// TIA Portal project "Øvelser_2_3_4_5_6_8" (V16)

(* hardware
DEVICE "S7-1200 station_1"  S7-1200 Station
   slot 0: "Rack_0"  S7-1200 Rack  Rack  V1.0
   slot 1: "PLC_1"  CPU 1214C DC/DC/DC  6ES7 214-1AG40-0XB0  V4.4
   slot 3: "AQ 1x12BIT_1"  AQ1 signal board  6ES7 232-4HA30-0XB0  V1.0
DEVICE "HMI_1"  KTP700 Basic PN
   slot 0: "HMI_1"  KTP700 Basic PN  6AV2 123-2GB03-0AX0  16.0.0.0
   slot 1: "HMI_RT_1"  KTP700 Basic PN  6AV2 123-2GB03-0AX0  16.0.0.0
   slot 5: "HMI_1.IE_CP_1"  PROFINET Interface  16.0.0.0
      slot 1: "PROFINET Interface_1"  PROFINET Interface
         slot 1: "Port_1"  Port
*)

// ===== PLC "PLC_1"  CPU 1214C DC/DC/DC =====

VAR_GLOBAL   // PLC tag table "Default tag table"
   "AutoHighCommand" AT %M2.0 : Bool;
   "TestStatus" AT %MW4 : Word;
   "HighCommand" AT %M2.1 : Bool;
   "LowCommand" AT %M2.2 : Bool;
   "SensorLow" AT %M2.4 : Bool;
   "IsHigh" AT %M2.5 : Bool;
   "IsLow" AT %M2.6 : Bool;
   "SensorIn" AT %I0.0 : Bool;
   "SensorOut" AT %I0.1 : Bool;
   "GoOut" AT %Q0.0 : Bool;
   "GoIn" AT %Q0.1 : Bool;
   "SensorUp" AT %I0.3 : Bool;
   "SensorDown" AT %I0.5 : Bool;
   "GoUp" AT %Q0.3 : Bool;
   "GoDown" AT %Q0.2 : Bool;
   "GrabCommand" AT %Q0.4 : Bool;
   "TestCommands" AT %MW0 : Word;
   "SensorHigh" AT %M2.3 : Bool;
   "IsIn" AT %M2.7 : Bool;
   "IsOut" AT %M3.0 : Bool;
   "AutoCommandGoOut" AT %M3.1 : Bool;
   "AutoCommandGoDown" AT %M3.2 : Bool;
   "AutoCommandGrab" AT %M3.3 : Bool;
   "IsUp" AT %M3.4 : Bool;
   "IsDown" AT %M3.5 : Bool;
   "HasGrapped" AT %M3.6 : Bool;
   "HasReleased" AT %M3.7 : Bool;
END_VAR

TYPE "TypeHMI_Commands"
   STRUCT
      Spare0 : Bool;   // (Bit 8), byteswap
      Spare1 : Bool;
      Spare2 : Bool;
      Spare3 : Bool;
      Spare4 : Bool;
      Spare5 : Bool;
      Spare6 : Bool;
      Spare7 : Bool;
      Manual : Bool;   // (Bit 0), byteswap
      Auto : Bool;
      ManualHighCommand : Bool;
      ManualLowCommand : Bool;
      SimulateFeddback : Bool;   // toggle simulation of feedback sensors
      Spare8 : Bool;
      Spare9 : Bool;
      Spare10 : Bool;
   END_STRUCT;
END_TYPE

TYPE "TypeHMI_Status"
   STRUCT
      AlarmToHigh : Bool;
      AlarmToLow : Bool;
      Spare2 : Bool;
      Spare3 : Bool;
      Spare4 : Bool;
      Spare5 : Bool;
      Spare6 : Bool;
      Spare7 : Bool;
      IsManual : Bool;
      IsHigh : Bool;
      IsLow : Bool;
      TransitionToHigh : Bool;
      TransitionToLow : Bool;
      FeedbackSensorLow : Bool;   // Satus, sensor
      FeedbackSensorHigh : Bool;   // Status, sensor
      FeedbackIsSimulated : Bool;
   END_STRUCT;
END_TYPE

DATA_BLOCK "Type_ControlModuleActuator_DB"   // DB1
{ S7_Optimized_Access := 'TRUE' }
VERSION : 0.1
// stored: InstanceOfName Type_ControlModuleActuator
"Type_ControlModuleActuator"
BEGIN
END_DATA_BLOCK

DATA_BLOCK "Type_ControlModuleActuator_DB_1"   // DB2
{ S7_Optimized_Access := 'TRUE' }
VERSION : 0.1
// stored: InstanceOfName Type_ControlModuleActuator
"Type_ControlModuleActuator"
BEGIN
END_DATA_BLOCK

DATA_BLOCK "Type_ControlModuleActuator_DB_2"   // DB3
{ S7_Optimized_Access := 'TRUE' }
VERSION : 0.1
// stored: InstanceOfName Type_ControlModuleActuator
"Type_ControlModuleActuator"
BEGIN
END_DATA_BLOCK

DATA_BLOCK "HMI"   // DB4
{ S7_Optimized_Access := 'TRUE' }
VERSION : 0.1
   VAR
      InOut : Struct
         Command : Word;
         Status : Word;
         StatusInt : Int;
      END_STRUCT;
      UpDown : Struct
         Command : Word;
         Status : Word;
         StatusInt : Int;
      END_STRUCT;
      Grab : Struct
         Command : Word;
         Status : Word;
         StatusInt : Int;
      END_STRUCT;
      TankCalculation : Struct
         CurrentLiguidLevel : Real;   // m
         Radius : Real;   // m
         ConeHight : Real;   // m
         Content : Real;   // m^3
      END_STRUCT;
      Sequence : Struct
         CommandAToB : Bool;
         CommandBToA : Bool;
         Status : Int;
      END_STRUCT;
   END_VAR
BEGIN
END_DATA_BLOCK

DATA_BLOCK "UpDown"   // DB5
{ S7_Optimized_Access := 'TRUE' }
VERSION : 0.1
// stored: InstanceOfName Type_ControlModuleActuator
"Type_ControlModuleActuator"
BEGIN
END_DATA_BLOCK

DATA_BLOCK "Grab"   // DB6
{ S7_Optimized_Access := 'TRUE' }
VERSION : 0.1
// stored: InstanceOfName Type_ControlModuleActuator
"Type_ControlModuleActuator"
BEGIN
END_DATA_BLOCK

DATA_BLOCK "HMI_alarms"   // DB9
{ S7_Optimized_Access := 'TRUE' }
VERSION : 0.1
   VAR
      alarm1 : Bool;
      alarm2 : Bool;
      alarm3 : Bool;
      alarm4 : Bool;
      alarm5 : Bool;
      alarm6 : Bool;
   END_VAR
BEGIN
END_DATA_BLOCK

DATA_BLOCK "Sequence_DB"   // DB10
{ S7_Optimized_Access := 'TRUE' }
VERSION : 0.1
// stored: InstanceOfName Sequence
"Sequence"
BEGIN
END_DATA_BLOCK

// folder: System blocks/Program resources

DATA_BLOCK "IEC_Timer_0_DB"   // DB7
{ S7_Optimized_Access := 'TRUE' }
AUTHOR : Simatic
FAMILY : IEC
NAME : IEC_TMR
VERSION : 1.0
// stored: InstanceOfName IEC_TIMER
"IEC_TIMER"
BEGIN
END_DATA_BLOCK

DATA_BLOCK "IEC_Timer_0_DB_1"   // DB8
{ S7_Optimized_Access := 'TRUE' }
AUTHOR : Simatic
FAMILY : IEC
NAME : IEC_TMR
VERSION : 1.0
// stored: InstanceOfName IEC_TIMER
"IEC_TIMER"
BEGIN
END_DATA_BLOCK

// folder: (top level)

FUNCTION_BLOCK "Type_ControlModuleActuator"   // FB1, LAD
{ S7_Optimized_Access := 'TRUE' }
VERSION : 0.1
   VAR_INPUT
      InHMICommands : Word;
      HMI_Commands AT InHMICommands : "TypeHMI_Commands";
      AutoHighCommand : Bool;
      FeedbackSensorHigh : Bool;
      FeedbackSensorLow : Bool;
      FeedbackTime : Time;
   END_VAR
   VAR_OUTPUT
      OutHMIStatus : Word;
      HMI_Status AT OutHMIStatus : "TypeHMI_Status";
      StatusInt : Int;
      HighCommand : Bool;
      LowCommand : Bool;
      IsHigh : Bool;
      IsLow : Bool;
   END_VAR
   VAR
      Manual : Bool;
      StaticHighCommand : Bool;
      StaticIsSimulated : Bool;
      SimulatedHigh : Bool;
      SimulatedLow : Bool;
      HighAlarmTimer : TON_TIME;
      LowAlarmTimer : TON_TIME;
   END_VAR
BEGIN

REGION Network 1: Manual/Auto
   // controlled by HMI
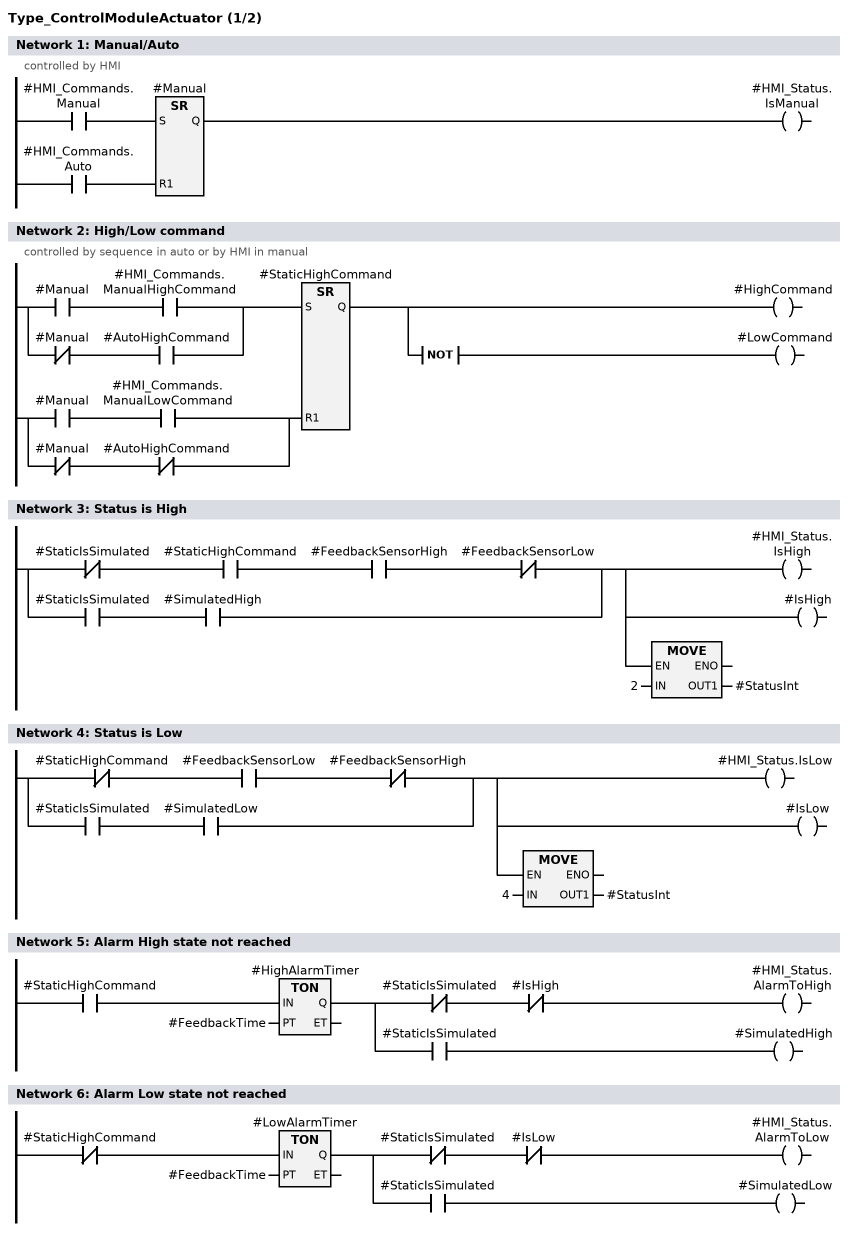
   RUNG wire#powerrail
      Contact( #HMI_Commands.Manual )
      S_SR(operand := #Manual, r1 := wire#w1)
      Coil( #HMI_Status.IsManual )
   END_RUNG
   RUNG wire#powerrail
      Contact( #HMI_Commands.Auto )
   END_RUNG wire#w1
   // the same network as SCL:
   IF #HMI_Commands.Manual THEN
       #Manual := TRUE;   // SR flip-flop
   END_IF;
   IF #HMI_Commands.Auto THEN #Manual := FALSE; END_IF;
   #HMI_Status.IsManual := #Manual;
END_REGION

REGION Network 2: High/Low command
   // controlled by sequence in auto or by HMI in manual
   RUNG wire#powerrail
      Contact( #Manual )
      Contact( #HMI_Commands.ManualHighCommand )
      wire#w1
      S_SR(operand := #StaticHighCommand, r1 := wire#w2)
      wire#w3
      Coil( #HighCommand )
   END_RUNG
   RUNG wire#powerrail
      I_Contact( #Manual )
      Contact( #AutoHighCommand )
   END_RUNG wire#w1
   RUNG wire#powerrail
      Contact( #Manual )
      Contact( #HMI_Commands.ManualLowCommand )
   END_RUNG wire#w2
   RUNG wire#powerrail
      I_Contact( #Manual )
      I_Contact( #AutoHighCommand )
   END_RUNG wire#w2
   RUNG wire#w3
      Not()
      Coil( #LowCommand )
   END_RUNG
   // the same network as SCL:
   IF (#Manual AND #HMI_Commands.ManualHighCommand) OR (NOT #Manual AND #AutoHighCommand) THEN
       #StaticHighCommand := TRUE;   // SR flip-flop
   END_IF;
   IF (#Manual AND #HMI_Commands.ManualLowCommand) OR (NOT #Manual AND NOT #AutoHighCommand) THEN
       #StaticHighCommand := FALSE;
   END_IF;
   #HighCommand := #StaticHighCommand;
   #LowCommand := NOT #StaticHighCommand;
END_REGION

REGION Network 3: Status is High
   RUNG wire#powerrail
      I_Contact( #StaticIsSimulated )
      Contact( #StaticHighCommand )
      Contact( #FeedbackSensorHigh )
      I_Contact( #FeedbackSensorLow )
      wire#w1
      Coil( #HMI_Status.IsHigh )
   END_RUNG
   RUNG wire#powerrail
      Contact( #StaticIsSimulated )
      Contact( #SimulatedHigh )
   END_RUNG wire#w1
   RUNG wire#w1
      Coil( #IsHigh )
   END_RUNG
   RUNG wire#w1
      Move(in := 2, out1 => #StatusInt)
   END_RUNG
   // the same network as SCL:
   #HMI_Status.IsHigh := (NOT #StaticIsSimulated AND #StaticHighCommand AND #FeedbackSensorHigh AND NOT #FeedbackSensorLow) OR (#StaticIsSimulated AND #SimulatedHigh);
   #IsHigh := #HMI_Status.IsHigh;
   IF #HMI_Status.IsHigh THEN #StatusInt := 2; END_IF;
END_REGION

REGION Network 4: Status is Low
   RUNG wire#powerrail
      I_Contact( #StaticHighCommand )
      Contact( #FeedbackSensorLow )
      I_Contact( #FeedbackSensorHigh )
      wire#w1
      Coil( #HMI_Status.IsLow )
   END_RUNG
   RUNG wire#powerrail
      Contact( #StaticIsSimulated )
      Contact( #SimulatedLow )
   END_RUNG wire#w1
   RUNG wire#w1
      Coil( #IsLow )
   END_RUNG
   RUNG wire#w1
      Move(in := 4, out1 => #StatusInt)
   END_RUNG
   // the same network as SCL:
   #HMI_Status.IsLow := (NOT #StaticHighCommand AND #FeedbackSensorLow AND NOT #FeedbackSensorHigh) OR (#StaticIsSimulated AND #SimulatedLow);
   #IsLow := #HMI_Status.IsLow;
   IF #HMI_Status.IsLow THEN #StatusInt := 4; END_IF;
END_REGION

REGION Network 5: Alarm High state not reached
   #HighAlarmTimer(IN := #StaticHighCommand, PT := #FeedbackTime);   // TON
   #HMI_Status.AlarmToHigh := #HighAlarmTimer.Q AND NOT #StaticIsSimulated AND NOT #IsHigh;
   #SimulatedHigh := #HighAlarmTimer.Q AND #StaticIsSimulated;
END_REGION

REGION Network 6: Alarm Low state not reached
   #LowAlarmTimer(IN := NOT #StaticHighCommand, PT := #FeedbackTime);   // TON
   #HMI_Status.AlarmToLow := #LowAlarmTimer.Q AND NOT #StaticIsSimulated AND NOT #IsLow;
   #SimulatedLow := #LowAlarmTimer.Q AND #StaticIsSimulated;
END_REGION

REGION Network 7: Togle simulation
END_REGION

REGION Network 8: Transition to High
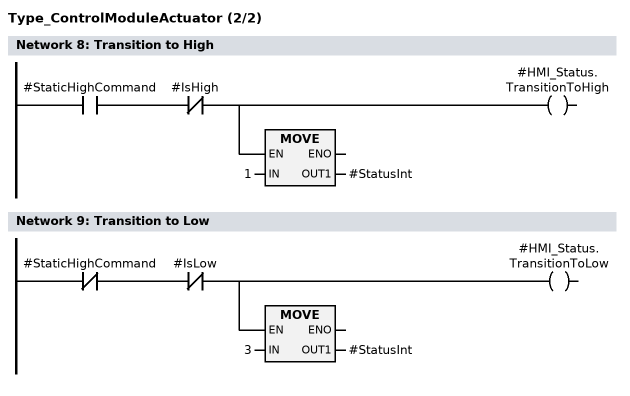
   RUNG wire#powerrail
      Contact( #StaticHighCommand )
      I_Contact( #IsHigh )
      wire#w1
      Coil( #HMI_Status.TransitionToHigh )
   END_RUNG
   RUNG wire#w1
      Move(in := 1, out1 => #StatusInt)
   END_RUNG
   // the same network as SCL:
   #HMI_Status.TransitionToHigh := #StaticHighCommand AND NOT #IsHigh;
   IF #HMI_Status.TransitionToHigh THEN #StatusInt := 1; END_IF;
END_REGION

REGION Network 9: Transition to Low
   RUNG wire#powerrail
      I_Contact( #StaticHighCommand )
      I_Contact( #IsLow )
      wire#w1
      Coil( #HMI_Status.TransitionToLow )
   END_RUNG
   RUNG wire#w1
      Move(in := 3, out1 => #StatusInt)
   END_RUNG
   // the same network as SCL:
   #HMI_Status.TransitionToLow := NOT #StaticHighCommand AND NOT #IsLow;
   IF #HMI_Status.TransitionToLow THEN #StatusInt := 3; END_IF;
END_REGION
END_FUNCTION_BLOCK

FUNCTION_BLOCK "Sequence"   // FB2, LAD
{ S7_Optimized_Access := 'TRUE' }
VERSION : 0.1
   VAR_INPUT
      AToB : Bool;
      BtoA : Bool;
      IsIn : Bool;
      IsOut : Bool;
      IsUp : Bool;
      IsDown : Bool;
      HasGrapped : Bool;
      HasReleased : Bool;
   END_VAR
   VAR_OUTPUT
      AutoCommandGoOut : Bool;
      AutoCommandGoDown : Bool;
      AutoCommandGrab : Bool;
      StatusStepNr : Int;
   END_VAR
   VAR
      StepNr : Int;
   END_VAR
   VAR_TEMP   // added for the SCL form of the ladder/FBD networks
      _w1 : Bool;
   END_VAR
BEGIN

REGION Network 1: Step 0:Idle
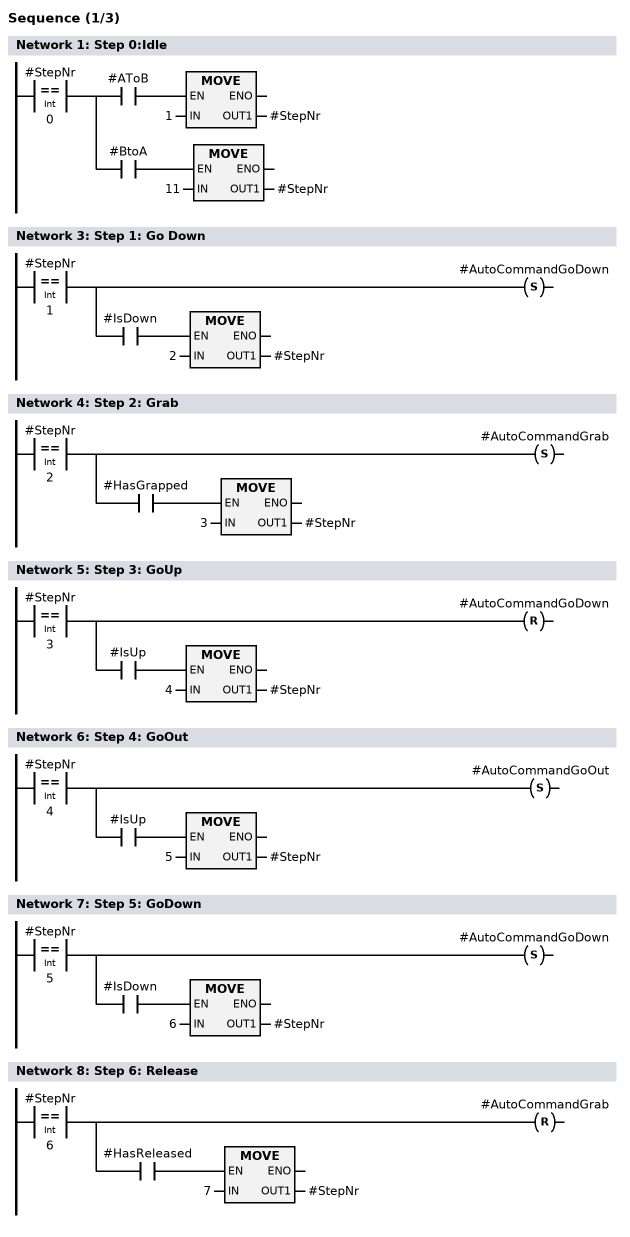
   RUNG wire#powerrail
      { S7_Templates := "SrcType := Int" } EQ_Contact(in1 := #StepNr, in2 := 0)
      wire#w1
      Contact( #AToB )
      Move(in := 1, out1 => #StepNr)
   END_RUNG
   RUNG wire#w1
      Contact( #BtoA )
      Move(in := 11, out1 => #StepNr)
   END_RUNG
   // the same network as SCL:
   #_w1 := #StepNr = 0;
   IF #_w1 AND #AToB THEN #StepNr := 1; END_IF;
   IF #_w1 AND #BtoA THEN #StepNr := 11; END_IF;
END_REGION

REGION Network 2: AToB
END_REGION

REGION Network 3: Step 1: Go Down
   RUNG wire#powerrail
      { S7_Templates := "SrcType := Int" } EQ_Contact(in1 := #StepNr, in2 := 1)
      wire#w1
      S_Coil( #AutoCommandGoDown )
   END_RUNG
   RUNG wire#w1
      Contact( #IsDown )
      Move(in := 2, out1 => #StepNr)
   END_RUNG
   // the same network as SCL:
   #_w1 := #StepNr = 1;
   IF #_w1 THEN #AutoCommandGoDown := TRUE; END_IF;
   IF #_w1 AND #IsDown THEN #StepNr := 2; END_IF;
END_REGION

REGION Network 4: Step 2: Grab
   RUNG wire#powerrail
      { S7_Templates := "SrcType := Int" } EQ_Contact(in1 := #StepNr, in2 := 2)
      wire#w1
      S_Coil( #AutoCommandGrab )
   END_RUNG
   RUNG wire#w1
      Contact( #HasGrapped )
      Move(in := 3, out1 => #StepNr)
   END_RUNG
   // the same network as SCL:
   #_w1 := #StepNr = 2;
   IF #_w1 THEN #AutoCommandGrab := TRUE; END_IF;
   IF #_w1 AND #HasGrapped THEN #StepNr := 3; END_IF;
END_REGION

REGION Network 5: Step 3: GoUp
   RUNG wire#powerrail
      { S7_Templates := "SrcType := Int" } EQ_Contact(in1 := #StepNr, in2 := 3)
      wire#w1
      R_Coil( #AutoCommandGoDown )
   END_RUNG
   RUNG wire#w1
      Contact( #IsUp )
      Move(in := 4, out1 => #StepNr)
   END_RUNG
   // the same network as SCL:
   #_w1 := #StepNr = 3;
   IF #_w1 THEN #AutoCommandGoDown := FALSE; END_IF;
   IF #_w1 AND #IsUp THEN #StepNr := 4; END_IF;
END_REGION

REGION Network 6: Step 4: GoOut
   RUNG wire#powerrail
      { S7_Templates := "SrcType := Int" } EQ_Contact(in1 := #StepNr, in2 := 4)
      wire#w1
      S_Coil( #AutoCommandGoOut )
   END_RUNG
   RUNG wire#w1
      Contact( #IsUp )
      Move(in := 5, out1 => #StepNr)
   END_RUNG
   // the same network as SCL:
   #_w1 := #StepNr = 4;
   IF #_w1 THEN #AutoCommandGoOut := TRUE; END_IF;
   IF #_w1 AND #IsUp THEN #StepNr := 5; END_IF;
END_REGION

REGION Network 7: Step 5: GoDown
   RUNG wire#powerrail
      { S7_Templates := "SrcType := Int" } EQ_Contact(in1 := #StepNr, in2 := 5)
      wire#w1
      S_Coil( #AutoCommandGoDown )
   END_RUNG
   RUNG wire#w1
      Contact( #IsDown )
      Move(in := 6, out1 => #StepNr)
   END_RUNG
   // the same network as SCL:
   #_w1 := #StepNr = 5;
   IF #_w1 THEN #AutoCommandGoDown := TRUE; END_IF;
   IF #_w1 AND #IsDown THEN #StepNr := 6; END_IF;
END_REGION

REGION Network 8: Step 6: Release
   RUNG wire#powerrail
      { S7_Templates := "SrcType := Int" } EQ_Contact(in1 := #StepNr, in2 := 6)
      wire#w1
      R_Coil( #AutoCommandGrab )
   END_RUNG
   RUNG wire#w1
      Contact( #HasReleased )
      Move(in := 7, out1 => #StepNr)
   END_RUNG
   // the same network as SCL:
   #_w1 := #StepNr = 6;
   IF #_w1 THEN #AutoCommandGrab := FALSE; END_IF;
   IF #_w1 AND #HasReleased THEN #StepNr := 7; END_IF;
END_REGION

REGION Network 9: Step 2: GoUp
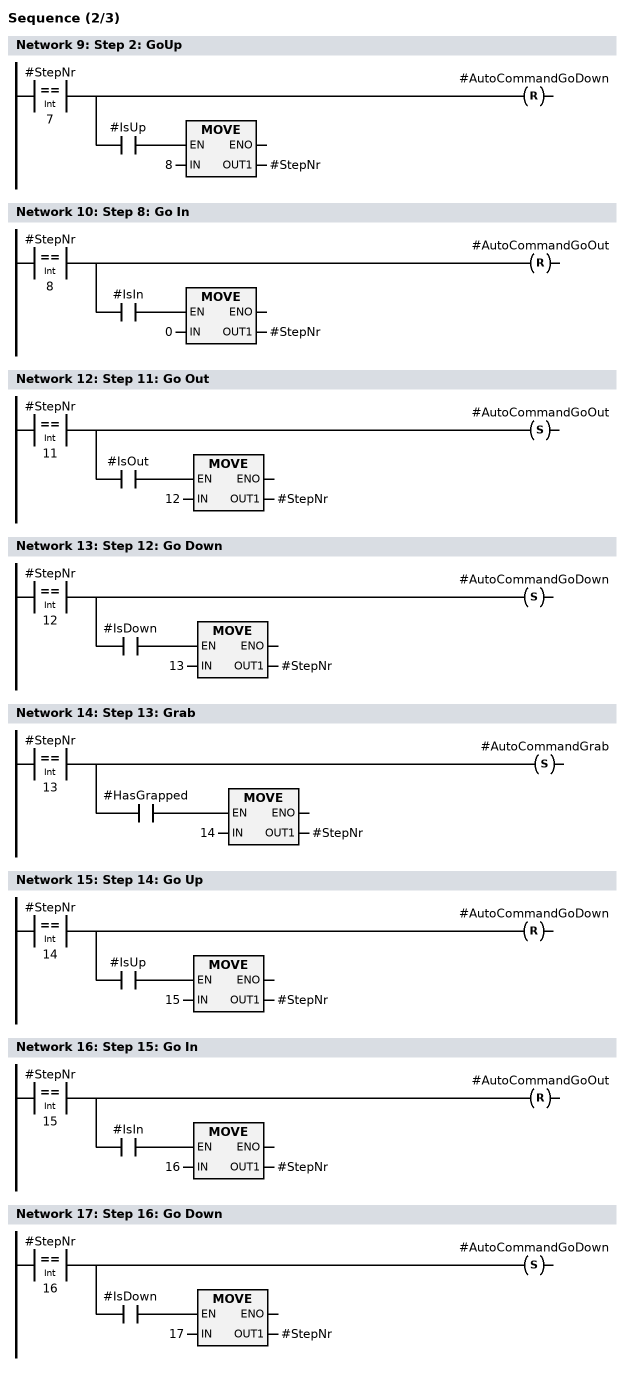
   RUNG wire#powerrail
      { S7_Templates := "SrcType := Int" } EQ_Contact(in1 := #StepNr, in2 := 7)
      wire#w1
      R_Coil( #AutoCommandGoDown )
   END_RUNG
   RUNG wire#w1
      Contact( #IsUp )
      Move(in := 8, out1 => #StepNr)
   END_RUNG
   // the same network as SCL:
   #_w1 := #StepNr = 7;
   IF #_w1 THEN #AutoCommandGoDown := FALSE; END_IF;
   IF #_w1 AND #IsUp THEN #StepNr := 8; END_IF;
END_REGION

REGION Network 10: Step 8: Go In
   RUNG wire#powerrail
      { S7_Templates := "SrcType := Int" } EQ_Contact(in1 := #StepNr, in2 := 8)
      wire#w1
      R_Coil( #AutoCommandGoOut )
   END_RUNG
   RUNG wire#w1
      Contact( #IsIn )
      Move(in := 0, out1 => #StepNr)
   END_RUNG
   // the same network as SCL:
   #_w1 := #StepNr = 8;
   IF #_w1 THEN #AutoCommandGoOut := FALSE; END_IF;
   IF #_w1 AND #IsIn THEN #StepNr := 0; END_IF;
END_REGION

REGION Network 11: BToA
END_REGION

REGION Network 12: Step 11: Go Out
   RUNG wire#powerrail
      { S7_Templates := "SrcType := Int" } EQ_Contact(in1 := #StepNr, in2 := 11)
      wire#w1
      S_Coil( #AutoCommandGoOut )
   END_RUNG
   RUNG wire#w1
      Contact( #IsOut )
      Move(in := 12, out1 => #StepNr)
   END_RUNG
   // the same network as SCL:
   #_w1 := #StepNr = 11;
   IF #_w1 THEN #AutoCommandGoOut := TRUE; END_IF;
   IF #_w1 AND #IsOut THEN #StepNr := 12; END_IF;
END_REGION

REGION Network 13: Step 12: Go Down
   RUNG wire#powerrail
      { S7_Templates := "SrcType := Int" } EQ_Contact(in1 := #StepNr, in2 := 12)
      wire#w1
      S_Coil( #AutoCommandGoDown )
   END_RUNG
   RUNG wire#w1
      Contact( #IsDown )
      Move(in := 13, out1 => #StepNr)
   END_RUNG
   // the same network as SCL:
   #_w1 := #StepNr = 12;
   IF #_w1 THEN #AutoCommandGoDown := TRUE; END_IF;
   IF #_w1 AND #IsDown THEN #StepNr := 13; END_IF;
END_REGION

REGION Network 14: Step 13: Grab
   RUNG wire#powerrail
      { S7_Templates := "SrcType := Int" } EQ_Contact(in1 := #StepNr, in2 := 13)
      wire#w1
      S_Coil( #AutoCommandGrab )
   END_RUNG
   RUNG wire#w1
      Contact( #HasGrapped )
      Move(in := 14, out1 => #StepNr)
   END_RUNG
   // the same network as SCL:
   #_w1 := #StepNr = 13;
   IF #_w1 THEN #AutoCommandGrab := TRUE; END_IF;
   IF #_w1 AND #HasGrapped THEN #StepNr := 14; END_IF;
END_REGION

REGION Network 15: Step 14: Go Up
   RUNG wire#powerrail
      { S7_Templates := "SrcType := Int" } EQ_Contact(in1 := #StepNr, in2 := 14)
      wire#w1
      R_Coil( #AutoCommandGoDown )
   END_RUNG
   RUNG wire#w1
      Contact( #IsUp )
      Move(in := 15, out1 => #StepNr)
   END_RUNG
   // the same network as SCL:
   #_w1 := #StepNr = 14;
   IF #_w1 THEN #AutoCommandGoDown := FALSE; END_IF;
   IF #_w1 AND #IsUp THEN #StepNr := 15; END_IF;
END_REGION

REGION Network 16: Step 15: Go In
   RUNG wire#powerrail
      { S7_Templates := "SrcType := Int" } EQ_Contact(in1 := #StepNr, in2 := 15)
      wire#w1
      R_Coil( #AutoCommandGoOut )
   END_RUNG
   RUNG wire#w1
      Contact( #IsIn )
      Move(in := 16, out1 => #StepNr)
   END_RUNG
   // the same network as SCL:
   #_w1 := #StepNr = 15;
   IF #_w1 THEN #AutoCommandGoOut := FALSE; END_IF;
   IF #_w1 AND #IsIn THEN #StepNr := 16; END_IF;
END_REGION

REGION Network 17: Step 16: Go Down
   RUNG wire#powerrail
      { S7_Templates := "SrcType := Int" } EQ_Contact(in1 := #StepNr, in2 := 16)
      wire#w1
      S_Coil( #AutoCommandGoDown )
   END_RUNG
   RUNG wire#w1
      Contact( #IsDown )
      Move(in := 17, out1 => #StepNr)
   END_RUNG
   // the same network as SCL:
   #_w1 := #StepNr = 16;
   IF #_w1 THEN #AutoCommandGoDown := TRUE; END_IF;
   IF #_w1 AND #IsDown THEN #StepNr := 17; END_IF;
END_REGION

REGION Network 18: Step 17: Release
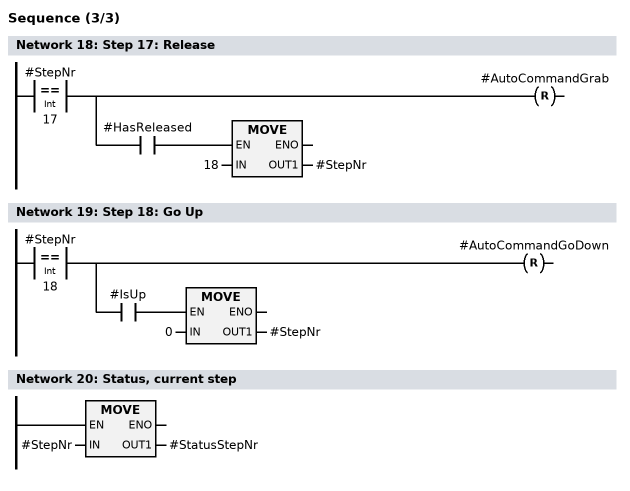
   RUNG wire#powerrail
      { S7_Templates := "SrcType := Int" } EQ_Contact(in1 := #StepNr, in2 := 17)
      wire#w1
      R_Coil( #AutoCommandGrab )
   END_RUNG
   RUNG wire#w1
      Contact( #HasReleased )
      Move(in := 18, out1 => #StepNr)
   END_RUNG
   // the same network as SCL:
   #_w1 := #StepNr = 17;
   IF #_w1 THEN #AutoCommandGrab := FALSE; END_IF;
   IF #_w1 AND #HasReleased THEN #StepNr := 18; END_IF;
END_REGION

REGION Network 19: Step 18: Go Up
   RUNG wire#powerrail
      { S7_Templates := "SrcType := Int" } EQ_Contact(in1 := #StepNr, in2 := 18)
      wire#w1
      R_Coil( #AutoCommandGoDown )
   END_RUNG
   RUNG wire#w1
      Contact( #IsUp )
      Move(in := 0, out1 => #StepNr)
   END_RUNG
   // the same network as SCL:
   #_w1 := #StepNr = 18;
   IF #_w1 THEN #AutoCommandGoDown := FALSE; END_IF;
   IF #_w1 AND #IsUp THEN #StepNr := 0; END_IF;
END_REGION

REGION Network 20: Status, current step
   RUNG wire#powerrail
      Move(in := #StepNr, out1 => #StatusStepNr)
   END_RUNG
   // the same network as SCL:
   #StatusStepNr := #StepNr;
END_REGION
END_FUNCTION_BLOCK

FUNCTION "Tankberegner" : Void   // FC1, LAD
{ S7_Optimized_Access := 'TRUE' }
VERSION : 0.1
   VAR_INPUT
      ActualLiguidLevel : Real;   // [m]
      TankRadius : Real;
      ConeHight : Real;
   END_VAR
   VAR_OUTPUT
      ActualContent : Real;   // [m^3]
   END_VAR
   VAR_TEMP
      VæskehojdeKegle : Real;
      VæskehojdeCylinder : Real;
      ForholdstalRadiusKegle : Real;
      IndholdKegle : Real;
      IndholdCylinder : Real;
   END_VAR
   VAR CONSTANT
      Pi : Real := 3.141593;
   END_VAR
   VAR_TEMP   // added for the SCL form of the ladder/FBD networks
      _w1 : Bool;
   END_VAR
BEGIN

REGION Network 1: Find væskehojden i keglen og væskehojden i cylinderen
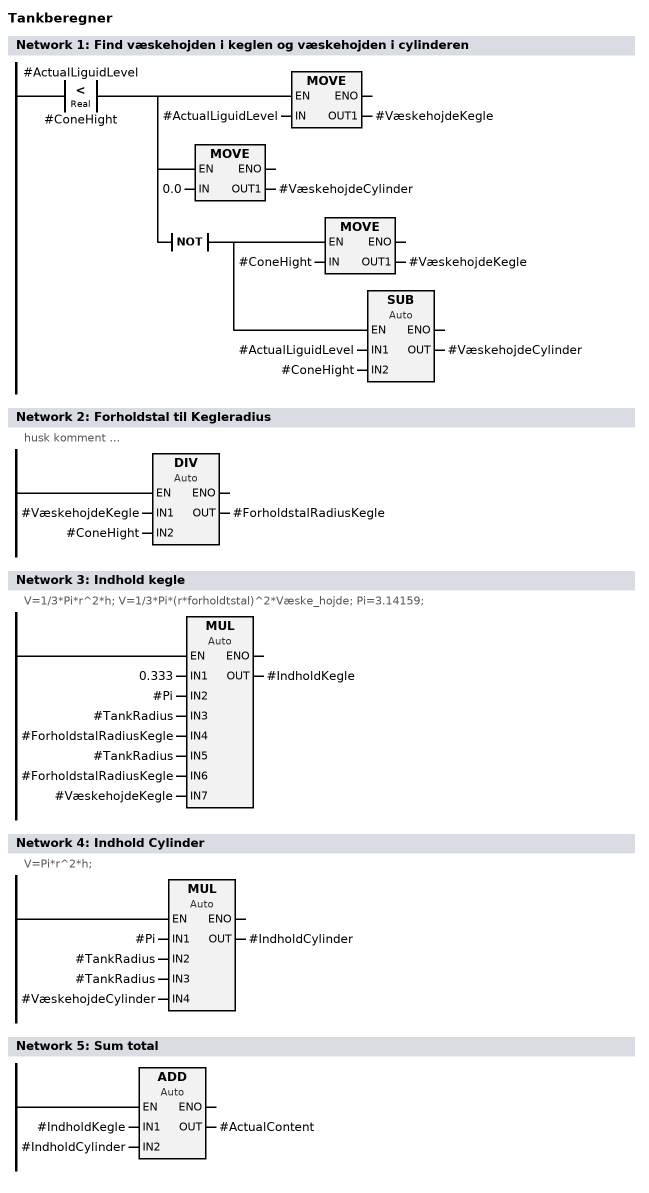
   RUNG wire#powerrail
      { S7_Templates := "SrcType := Real" } LT_Contact(in1 := #ActualLiguidLevel, in2 := #ConeHight)
      wire#w1
      Move(in := #ActualLiguidLevel, out1 => #VæskehojdeKegle)
   END_RUNG
   RUNG wire#w1
      Move(in := 0.0, out1 => #VæskehojdeCylinder)
   END_RUNG
   RUNG wire#w1
      Not()
      wire#w2
      Move(in := #ConeHight, out1 => #VæskehojdeKegle)
   END_RUNG
   RUNG wire#w2
      Sub(in1 := #ActualLiguidLevel, in2 := #ConeHight, out => #VæskehojdeCylinder)
   END_RUNG
   // the same network as SCL:
   #_w1 := #ActualLiguidLevel < #ConeHight;
   IF #_w1 THEN
       #VæskehojdeKegle := #ActualLiguidLevel;
       #VæskehojdeCylinder := 0.0;
   END_IF;
   IF NOT #_w1 THEN
       #VæskehojdeKegle := #ConeHight;
       #VæskehojdeCylinder := #ActualLiguidLevel - #ConeHight;
   END_IF;
END_REGION

REGION Network 2: Forholdstal til Kegleradius
   // husk komment ...
   RUNG wire#powerrail
      Div(in1 := #VæskehojdeKegle, in2 := #ConeHight, out => #ForholdstalRadiusKegle)
   END_RUNG
   // the same network as SCL:
   #ForholdstalRadiusKegle := #VæskehojdeKegle / #ConeHight;
END_REGION

REGION Network 3: Indhold kegle
   // V=1/3*Pi*r^2*h; V=1/3*Pi*(r*forholdtstal)^2*Væske_hojde; Pi=3.14159;
   RUNG wire#powerrail
      Mul(in1 := 0.333, in2 := #Pi, in3 := #TankRadius, in4 := #ForholdstalRadiusKegle, in5 := #TankRadius, in6 := #ForholdstalRadiusKegle, in7 := #VæskehojdeKegle, out => #IndholdKegle)
   END_RUNG
   // the same network as SCL:
   #IndholdKegle := 0.333 * #Pi * #TankRadius * #ForholdstalRadiusKegle * #TankRadius * #ForholdstalRadiusKegle * #VæskehojdeKegle;
END_REGION

REGION Network 4: Indhold Cylinder
   // V=Pi*r^2*h;
   RUNG wire#powerrail
      Mul(in1 := #Pi, in2 := #TankRadius, in3 := #TankRadius, in4 := #VæskehojdeCylinder, out => #IndholdCylinder)
   END_RUNG
   // the same network as SCL:
   #IndholdCylinder := #Pi * #TankRadius * #TankRadius * #VæskehojdeCylinder;
END_REGION

REGION Network 5: Sum total
   RUNG wire#powerrail
      Add(in1 := #IndholdKegle, in2 := #IndholdCylinder, out => #ActualContent)
   END_RUNG
   // the same network as SCL:
   #ActualContent := #IndholdKegle + #IndholdCylinder;
END_REGION
END_FUNCTION

ORGANIZATION_BLOCK "Main"   // OB1, LAD, ProgramCycle
TITLE = "Main Program Sweep (Cycle)"
{ S7_Optimized_Access := 'TRUE' }
VERSION : 0.1
   VAR_INPUT
      Initial_Call : Bool;   // Initial call of this OB
      Remanence : Bool;   // =True, if remanent data are available
   END_VAR
BEGIN

REGION Network 1: In/Out control modul
   // High=Out
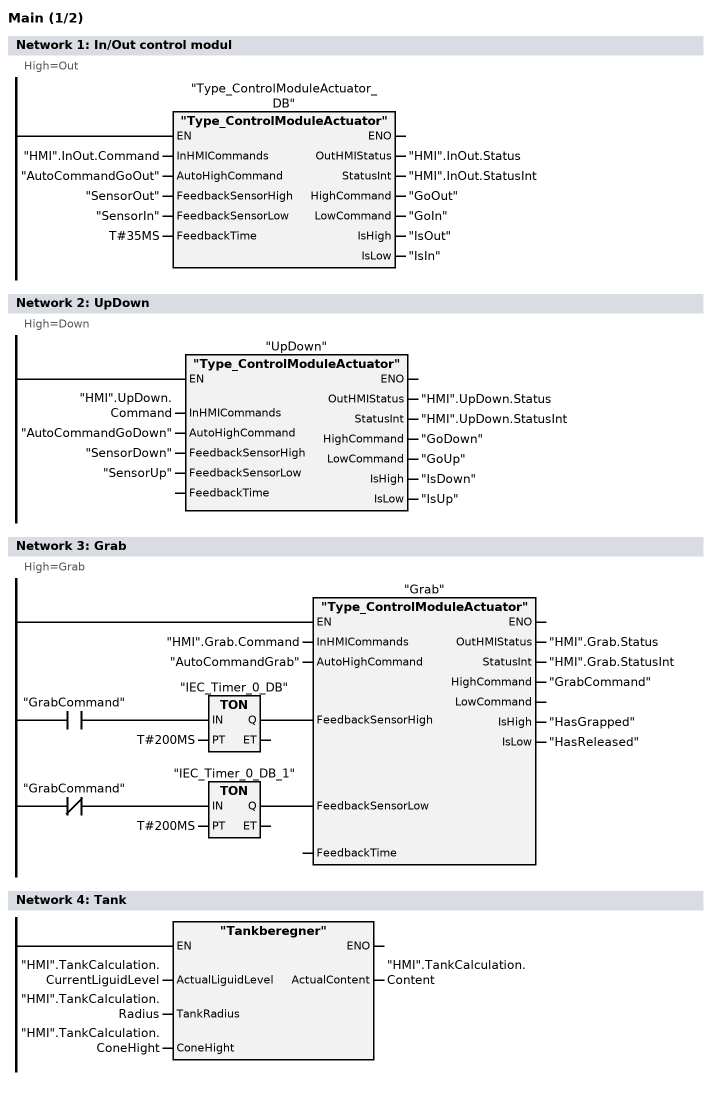
   RUNG wire#powerrail
      "Type_ControlModuleActuator_DB"(InHMICommands := "HMI".InOut.Command, AutoHighCommand := "AutoCommandGoOut", FeedbackSensorHigh := "SensorOut", FeedbackSensorLow := "SensorIn", FeedbackTime := T#35MS, OutHMIStatus => "HMI".InOut.Status, StatusInt => "HMI".InOut.StatusInt, HighCommand => "GoOut", LowCommand => "GoIn", IsHigh => "IsOut", IsLow => "IsIn")
   END_RUNG
   // the same network as SCL:
   "Type_ControlModuleActuator_DB"(InHMICommands := "HMI".InOut.Command,   // "Type_ControlModuleActuator"
                           AutoHighCommand := "AutoCommandGoOut",
                           FeedbackSensorHigh := "SensorOut",
                           FeedbackSensorLow := "SensorIn",
                           FeedbackTime := T#35MS,
                           OutHMIStatus => "HMI".InOut.Status,
                           StatusInt => "HMI".InOut.StatusInt,
                           HighCommand => "GoOut",
                           LowCommand => "GoIn",
                           IsHigh => "IsOut",
                           IsLow => "IsIn");
END_REGION

REGION Network 2: UpDown
   // High=Down
   RUNG wire#powerrail
      "UpDown"(InHMICommands := "HMI".UpDown.Command, AutoHighCommand := "AutoCommandGoDown", FeedbackSensorHigh := "SensorDown", FeedbackSensorLow := "SensorUp", FeedbackTime :=, OutHMIStatus => "HMI".UpDown.Status, StatusInt => "HMI".UpDown.StatusInt, HighCommand => "GoDown", LowCommand => "GoUp", IsHigh => "IsDown", IsLow => "IsUp")
   END_RUNG
   // the same network as SCL:
   "UpDown"(InHMICommands := "HMI".UpDown.Command,   // "Type_ControlModuleActuator"
            AutoHighCommand := "AutoCommandGoDown",
            FeedbackSensorHigh := "SensorDown",
            FeedbackSensorLow := "SensorUp",
            OutHMIStatus => "HMI".UpDown.Status,
            StatusInt => "HMI".UpDown.StatusInt,
            HighCommand => "GoDown",
            LowCommand => "GoUp",
            IsHigh => "IsDown",
            IsLow => "IsUp");
END_REGION

REGION Network 3: Grab
   // High=Grab
   "IEC_Timer_0_DB".TON(IN := "GrabCommand", PT := T#200MS);
   "IEC_Timer_0_DB_1".TON(IN := NOT "GrabCommand", PT := T#200MS);
   "Grab"(InHMICommands := "HMI".Grab.Command,   // "Type_ControlModuleActuator"
          AutoHighCommand := "AutoCommandGrab",
          FeedbackSensorHigh := "IEC_Timer_0_DB".Q,
          FeedbackSensorLow := "IEC_Timer_0_DB_1".Q,
          OutHMIStatus => "HMI".Grab.Status,
          StatusInt => "HMI".Grab.StatusInt,
          HighCommand => "GrabCommand",
          IsHigh => "HasGrapped",
          IsLow => "HasReleased");
END_REGION

REGION Network 4: Tank
   RUNG wire#powerrail
      "Tankberegner"(ActualLiguidLevel := "HMI".TankCalculation.CurrentLiguidLevel, TankRadius := "HMI".TankCalculation.Radius, ConeHight := "HMI".TankCalculation.ConeHight, ActualContent => "HMI".TankCalculation.Content)
   END_RUNG
   // the same network as SCL:
   "Tankberegner"(ActualLiguidLevel := "HMI".TankCalculation.CurrentLiguidLevel,
                  TankRadius := "HMI".TankCalculation.Radius,
                  ConeHight := "HMI".TankCalculation.ConeHight,
                  ActualContent => "HMI".TankCalculation.Content);
END_REGION

REGION Network 5: Sequence
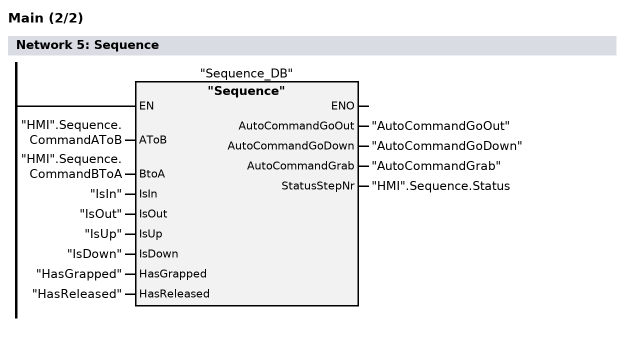
   RUNG wire#powerrail
      "Sequence_DB"(AToB := "HMI".Sequence.CommandAToB, BtoA := "HMI".Sequence.CommandBToA, IsIn := "IsIn", IsOut := "IsOut", IsUp := "IsUp", IsDown := "IsDown", HasGrapped := "HasGrapped", HasReleased := "HasReleased", AutoCommandGoOut => "AutoCommandGoOut", AutoCommandGoDown => "AutoCommandGoDown", AutoCommandGrab => "AutoCommandGrab", StatusStepNr => "HMI".Sequence.Status)
   END_RUNG
   // the same network as SCL:
   "Sequence_DB"(AToB := "HMI".Sequence.CommandAToB,   // "Sequence"
                 BtoA := "HMI".Sequence.CommandBToA,
                 IsIn := "IsIn",
                 IsOut := "IsOut",
                 IsUp := "IsUp",
                 IsDown := "IsDown",
                 HasGrapped := "HasGrapped",
                 HasReleased := "HasReleased",
                 AutoCommandGoOut => "AutoCommandGoOut",
                 AutoCommandGoDown => "AutoCommandGoDown",
                 AutoCommandGrab => "AutoCommandGrab",
                 StatusStepNr => "HMI".Sequence.Status);
END_REGION
END_ORGANIZATION_BLOCK

(* ===== HMI "HMI_RT_1" =====
system functions are stored by id; their names below are inferred from use
connection "HMI_Connection_1": ETHERNET, SMART_S7_1200_OMS

HMI tags "Default tag table"
   "HMI_InOut_Command" : Word = PLC HMI.InOut.Command, 1 s
   "HMI_InOut_Status" : Word = PLC HMI.InOut.Status, 1 s
   "HMI_UpDown_Command" : Word = PLC HMI.UpDown.Command, 1 s
   "HMI_UpDown_Status" : Word = PLC HMI.UpDown.Status, 1 s
   "HMI_Grab_Command" : Word = PLC HMI.Grab.Command, 1 s
   "HMI_Grab_Status" : Word = PLC HMI.Grab.Status, 1 s
   "HMI_InOut_StatusInt" : Int = PLC HMI.InOut.StatusInt, 1 s
   "HMI_UpDown_StatusInt" : Int = PLC HMI.UpDown.StatusInt, 1 s
   "HMI_Grab_StatusInt" : Int = PLC HMI.Grab.StatusInt, 1 s
   "HMI_TankCalculation_Radius" : Real = PLC HMI.TankCalculation.Radius, 1 s
   "HMI_TankCalculation_ConeHight" : Real = PLC HMI.TankCalculation.ConeHight, 1 s
   "HMI_TankCalculation_CurentLiguidLevel" : Real = PLC HMI.TankCalculation.CurrentLiguidLevel, 1 s
   "HMI_TankCalculation_Content" : Real = PLC HMI.TankCalculation.Content, 1 s
   "HMI_Sequence_CommandAToB" : Bool = PLC HMI.Sequence.CommandAToB, 1 s
   "HMI_Sequence_CommandBToA" : Bool = PLC HMI.Sequence.CommandBToA, 1 s

discrete alarms
   1: 'failed on the way out', class Errors, trigger "HMI_InOut_Status" bit 8
   2: 'failed on the way in', class Errors, trigger "HMI_InOut_Status" bit 9
   3: 'failed on the way down', class Errors, trigger "HMI_UpDown_Status" bit 8
   4: 'failed on the way up', class Errors, trigger "HMI_UpDown_Status" bit 9
   5: 'failed grab', class Errors, trigger "HMI_Grab_Status" bit 8
   6: 'failed reliease', class Errors, trigger "HMI_Grab_Status" bit 9

text list "upDown": 1 'GoingDown'; 2 'IsDown'; 3 'GoingUp'; 4 'IsUp'

text list "InOut": 1 'TransitionToOut'; 2 'IsOut'; 3 'TransitionToIn'; 4 'IsIn'

text list "Grab": 1 'Gripping'; 2 'Grabbed'; 3 'Releasing'; 4 'Released'

screen "InOut" 800x480
   Button "Button_1" at 73,290 size 96x32; TextOff 'Simulate'
      on Press: function_b14e0dd5("HMI_InOut_Command", 4)
   Button "Button_2" at 71,52 size 96x32; TextOff 'Manual'
      on Press: function_b14e0dd5("HMI_InOut_Command", 0)
   Button "Button_3" at 73,230 size 96x32; TextOff 'ManLow'
      on Press: function_b14e0dd5("HMI_InOut_Command", 3)
   Button "Button_4" at 73,171 size 96x32; TextOff 'ManHigh'
      on Press: function_b14e0dd5("HMI_InOut_Command", 2)
   Button "Button_6" at 73,111 size 96x32; TextOff 'Auto'
      on Press: function_b14e0dd5("HMI_InOut_Command", 1)
   Circle "Circle_1" at 185,52 size 34x34
      Appearance <- "HMI_InOut_Status"
   Circle "Circle_2" at 185,169 size 34x34
      Appearance <- "HMI_InOut_Status"
   Circle "Circle_3" at 185,225 size 34x34
      Appearance <- "HMI_InOut_Status"
   Circle "Circle_4" at 185,288 size 34x34
      Appearance <- "HMI_InOut_Status"
   TextField "Text field_1" at 367,30 size 51x23; Text 'InOut'
   Circle "Circle_5" at 238,168 size 34x34
      Appearance <- "HMI_InOut_Status"
   Circle "Circle_6" at 238,227 size 34x34
      Appearance <- "HMI_InOut_Status"

screen "Grab" 800x480
   Button "Button_1" at 73,290 size 96x32; TextOff 'Simulate'
      on Press: function_b14e0dd5("HMI_Grab_Command", 4)
   Button "Button_2" at 71,52 size 96x32; TextOff 'Manual'
      on Press: function_b14e0dd5("HMI_Grab_Command", 0)
   Button "Button_3" at 73,230 size 96x32; TextOff 'ManLow'
      on Press: function_b14e0dd5("HMI_Grab_Command", 3)
   Button "Button_4" at 73,171 size 96x32; TextOff 'ManHigh'
      on Press: function_b14e0dd5("HMI_Grab_Command", 2)
   Button "Button_6" at 73,111 size 96x32; TextOff 'Auto'
      on Press: function_b14e0dd5("HMI_Grab_Command", 1)
   Circle "Circle_1" at 185,52 size 34x34
      Appearance <- "HMI_Grab_Status"
   Circle "Circle_2" at 185,169 size 34x34
      Appearance <- "HMI_Grab_Status"
   Circle "Circle_3" at 185,225 size 34x34
      Appearance <- "HMI_Grab_Status"
   Circle "Circle_4" at 185,288 size 34x34
      Appearance <- "HMI_Grab_Status"
   TextField "Text field_1" at 367,30 size 44x23; Text 'Grab'
   Circle "Circle_5" at 238,168 size 34x34
      Appearance <- "HMI_Grab_Status"
   Circle "Circle_6" at 238,227 size 34x34
      Appearance <- "HMI_Grab_Status"

screen "UpDown" 800x480
   Button "Button_1" at 73,290 size 96x32; TextOff 'Simulate'
      on Press: function_b14e0dd5("HMI_UpDown_Command", 4)
   Button "Button_2" at 71,52 size 96x32; TextOff 'Manual'
      on Press: function_b14e0dd5("HMI_UpDown_Command", 0)
   Button "Button_3" at 73,230 size 96x32; TextOff 'ManLow'
      on Press: function_b14e0dd5("HMI_UpDown_Command", 3)
   Button "Button_4" at 73,171 size 96x32; TextOff 'ManHigh'
      on Press: function_b14e0dd5("HMI_UpDown_Command", 2)
   Button "Button_6" at 73,111 size 96x32; TextOff 'Auto'
      on Press: function_b14e0dd5("HMI_UpDown_Command", 1)
   Circle "Circle_1" at 185,52 size 34x34
      Appearance <- "HMI_UpDown_Status"
   Circle "Circle_2" at 185,169 size 34x34
      Appearance <- "HMI_UpDown_Status"
   Circle "Circle_3" at 185,225 size 34x34
      Appearance <- "HMI_UpDown_Status"
   Circle "Circle_4" at 185,288 size 34x34
      Appearance <- "HMI_UpDown_Status"
   TextField "Text field_1" at 367,30 size 73x23; Text 'UpDown'
   Circle "Circle_5" at 238,168 size 34x34
      Appearance <- "HMI_UpDown_Status"
   Circle "Circle_6" at 238,227 size 34x34
      Appearance <- "HMI_UpDown_Status"

screen "Home" 800x480
   SymbolicIOField "Symbolic I/O field_1" at 204,43 size 159x32; TextOn '1'; TextOff '0'; TextList "InOut"
      ProcessValue <- "HMI_InOut_StatusInt"
   TextField "Text field_1" at 45,40 size 108x23; Text 'InOut Status'
   SymbolicIOField "Symbolic I/O field_2" at 204,93 size 159x32; TextOn '1'; TextOff '0'; TextList "upDown"
      ProcessValue <- "HMI_UpDown_StatusInt"
   SymbolicIOField "Symbolic I/O field_3" at 204,143 size 159x32; TextOn '1'; TextOff '0'; TextList "Grab"
      ProcessValue <- "HMI_Grab_StatusInt"
   TextField "Text field_2" at 45,90 size 130x23; Text 'UpDown Status'
   TextField "Text field_3" at 49,143 size 94x23; Text 'Grab Satus'
   TextField "Text field_4" at 50,296 size 140x23; Text 'Sequence Status'
   Button "Button_1" at 228,284 size 96x32; TextOff 'AtoB'
      on Press: function_b14e0dd5("HMI_Sequence_CommandAToB", 0)
   Button "Button_2" at 359,287 size 96x32; TextOff 'BToA'
      on Press: function_b14e0dd5("HMI_Sequence_CommandBToA", 0)
   IOField "I/O field_1" at 228,351 size 96x32; FormatPattern 9999999
   IOField "I/O field_2" at 359,350 size 96x32; FormatPattern 9999999

screen "TankC" 800x480
   TextField "Text field_1" at 244,57 size 65x23; Text 'Radius'
   TextField "Text field_2" at 244,135 size 90x23; Text 'ConeHight'
   TextField "Text field_3" at 244,213 size 174x23; Text 'Current Liguid Level'
   TextField "Text field_4" at 244,292 size 75x23; Text 'Content'
   Bar "Bar_1" at 566,135 size 80x120; MinimumValue 0; MaximumValue 100
      ProcessValue <- "HMI_TankCalculation_Content"
   IOField "I/O field_1" at 39,48 size 96x32; FormatPattern s999999999.999
      ProcessValue <- "HMI_TankCalculation_Radius"
   IOField "I/O field_2" at 38,212 size 96x32; FormatPattern s999999999.999
      ProcessValue <- "HMI_TankCalculation_CurentLiguidLevel"
   IOField "I/O field_3" at 39,130 size 96x32; FormatPattern s999999999.999
      ProcessValue <- "HMI_TankCalculation_ConeHight"
   IOField "I/O field_4" at 39,295 size 96x32; FormatPattern s999999999.999
      ProcessValue <- "HMI_TankCalculation_Content"

screen "Alarm View" 800x480
   AlarmView "Alarm view_1" at 35,37 size 600x300
*)